(* Logix 5000 project; controller NWGG 1756-L72 rev 35.12; software revision 35.00; part 2 of 19 *)
(* tags used below, declared in another part *)
   T22 : TIMER[100];
   T4 : TIMER[100];

ADD_ON_INSTRUCTION Loadout_K_Valve_Control   (* revision 1.0 *)
VAR_IN_OUT
   K_Valve : udt_Loadout_K_Valve; {required}
   ALM_Clean_Pos_Failed : ALARM_DIGITAL; {required}
   ALM_Treat_Pos_Failed : ALARM_DIGITAL; {required}
   Treat_Position_Input : BOOL; {required}
   Clean_Position_Input : BOOL; {required}
   Clean_Gate_Relay : BOOL; {required}
   Treat_Gate_Relay : BOOL; {required}
END_VAR
VAR
   Clean_Pos_Failed_ACK : BOOL; {access None}
   Treat_Pos_Failedt_ACK : BOOL; {access None}
END_VAR

ROUTINE Logic   (* ladder *)
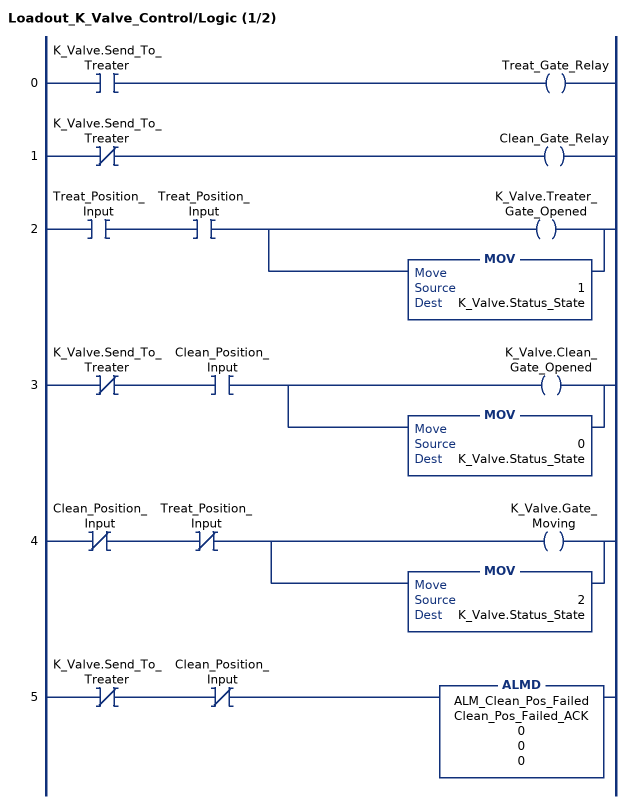
   0: XIC(K_Valve.Send_To_Treater)OTE(Treat_Gate_Relay);
   1: XIO(K_Valve.Send_To_Treater)OTE(Clean_Gate_Relay);
   2: XIC(Treat_Position_Input)XIC(Treat_Position_Input)[OTE(K_Valve.Treater_Gate_Opened) ,MOV(1,K_Valve.Status_State) ];
   3: XIO(K_Valve.Send_To_Treater)XIC(Clean_Position_Input)[OTE(K_Valve.Clean_Gate_Opened) ,MOV(0,K_Valve.Status_State) ];
   4: XIO(Clean_Position_Input)XIO(Treat_Position_Input)[OTE(K_Valve.Gate_Moving) ,MOV(2,K_Valve.Status_State) ];
   5: XIO(K_Valve.Send_To_Treater)XIO(Clean_Position_Input)ALMD(ALM_Clean_Pos_Failed,Clean_Pos_Failed_ACK,0,0,0);
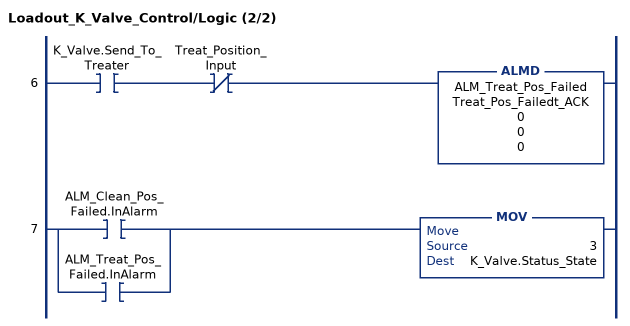
   6: XIC(K_Valve.Send_To_Treater)XIO(Treat_Position_Input)ALMD(ALM_Treat_Pos_Failed,Treat_Pos_Failedt_ACK,0,0,0);
   7: [XIC(ALM_Clean_Pos_Failed.InAlarm) ,XIC(ALM_Treat_Pos_Failed.InAlarm) ]MOV(3,K_Valve.Status_State);
END_ROUTINE
END_ADD_ON_INSTRUCTION

ADD_ON_INSTRUCTION Motor_Control   (* revision 1.0 *)
VAR_IN_OUT
   Motor_Contact : BOOL; {required}
END_VAR
VAR_INPUT
   Spd_20_Pct : BOOL; {required}
   Spd_10_Pct : BOOL; {required}
END_VAR
VAR_OUTPUT
   Running : BOOL; {access Read Only, required}
END_VAR
VAR_IN_OUT
   Motor_Alarm_SPD20 : ALARM_DIGITAL; {required}
   Motor_Alarm_SPD10 : ALARM_DIGITAL; {required}
   Motor_Alarm_Stopped_Over_Amps : ALARM_DIGITAL; {required}
   Motor_Start : udt_Motor_Start; {required}
END_VAR
VAR_INPUT
   Plugged_Sensor : BOOL; {required}
END_VAR
VAR_IN_OUT
   Motor_Alarm_Plugged : ALARM_DIGITAL; {required}
END_VAR
VAR_INPUT
   Motor_Amps : REAL; {required}
END_VAR
VAR_IN_OUT
   Motor_Config : udt_Motor_Config; {required}
   Motor_Starting : BOOL; {required}
   Motor_Alarm_Wont_Start : ALARM_DIGITAL; {required}
END_VAR
VAR_OUTPUT
   In_Alarm : BOOL; {access Read Only}
END_VAR
VAR_IN_OUT
   Treat_Batch_Status : DINT; {required}
   Clean_Batch_Status : DINT; {required}
   Transfer_Batch_Status : DINT; {required}
END_VAR
VAR_OUTPUT
   Motor_Batch_Ready : BOOL; {access Read Only}
END_VAR
VAR_IN_OUT
   Manual_Mode : BOOL; {required}
   InterLocked_Belt : BOOL; {required}
END_VAR
VAR_OUTPUT
   Motor_Batch_Ready_Clean : BOOL; {access Read Only}
   Motor_Batch_Ready_Treat : BOOL; {access Read Only}
   Motor_Batch_Ready_Transfer : BOOL; {access Read Only}
END_VAR
VAR
   TMR_BELT_SPD20 : TIMER := (PRE := 2000); {access None}
   TMR_AMP_INRUSH : TIMER := (PRE := 2000); {access None}
   Alm_Spd20_AK : BOOL; {access None}
   Alm_Spd10_AK : BOOL; {access None}
   Alm_Plugged_AK : BOOL; {access None}
   Alm_OVR_AMP_AK : BOOL; {access None}
   Stop_Motor_Plugged : BOOL; {access None}
   Stop_Motor_SLP20 : BOOL; {access None}
   Stop_Motor : BOOL; {access None}
   Stop_Motor_Ovr_Amp : BOOL; {access None}
   TMR_BELT_SPD10 : TIMER := (PRE := 2000); {access None}
   Alm_Wont_Start_AK : BOOL; {access None}
   Req_Motor_Start : BOOL; {access None}
   tmr_Auto_Stop_Delay : TIMER; {access None}
END_VAR

ROUTINE Logic   (* ladder *)
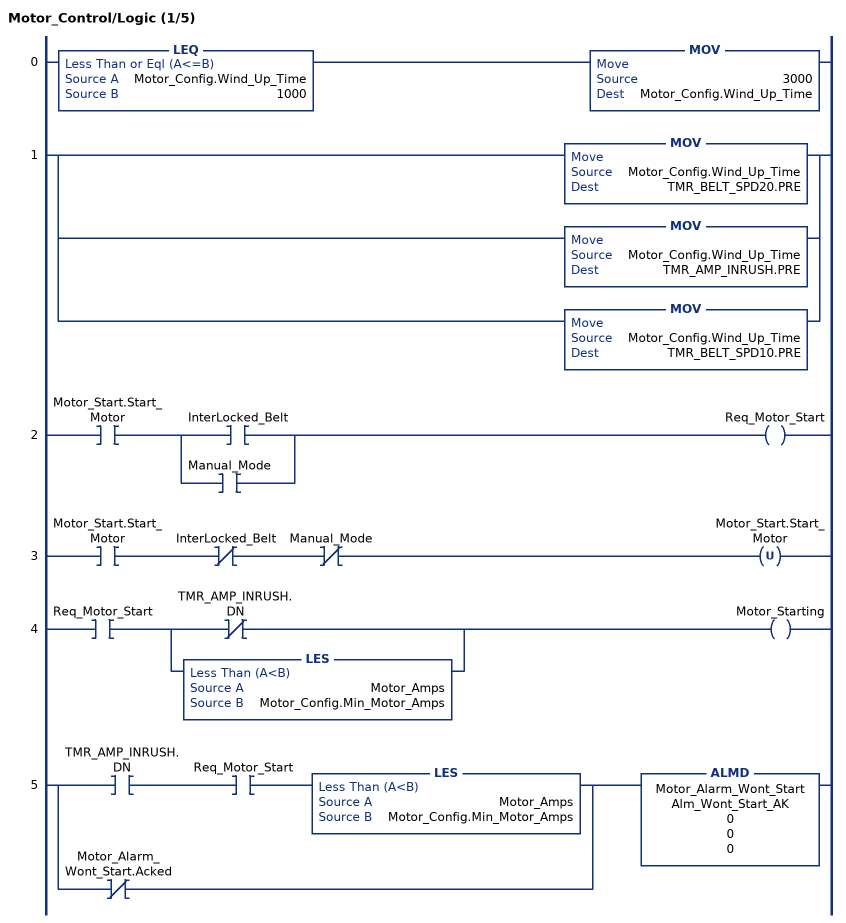
   0: LEQ(Motor_Config.Wind_Up_Time,1000)MOV(3000,Motor_Config.Wind_Up_Time);
   1: [MOV(Motor_Config.Wind_Up_Time,TMR_BELT_SPD20.PRE) ,MOV(Motor_Config.Wind_Up_Time,TMR_AMP_INRUSH.PRE) ,MOV(Motor_Config.Wind_Up_Time,TMR_BELT_SPD10.PRE) ];
   2: XIC(Motor_Start.Start_Motor)[XIC(InterLocked_Belt) ,XIC(Manual_Mode) ]OTE(Req_Motor_Start);
   3: XIC(Motor_Start.Start_Motor)XIO(InterLocked_Belt)XIO(Manual_Mode)OTU(Motor_Start.Start_Motor);
   4: XIC(Req_Motor_Start)[XIO(TMR_AMP_INRUSH.DN) ,LES(Motor_Amps,Motor_Config.Min_Motor_Amps) ]OTE(Motor_Starting);
   5: [XIC(TMR_AMP_INRUSH.DN) XIC(Req_Motor_Start) LES(Motor_Amps,Motor_Config.Min_Motor_Amps) ,XIO(Motor_Alarm_Wont_Start.Acked) ]ALMD(Motor_Alarm_Wont_Start,Alm_Wont_Start_AK,0,0,0);
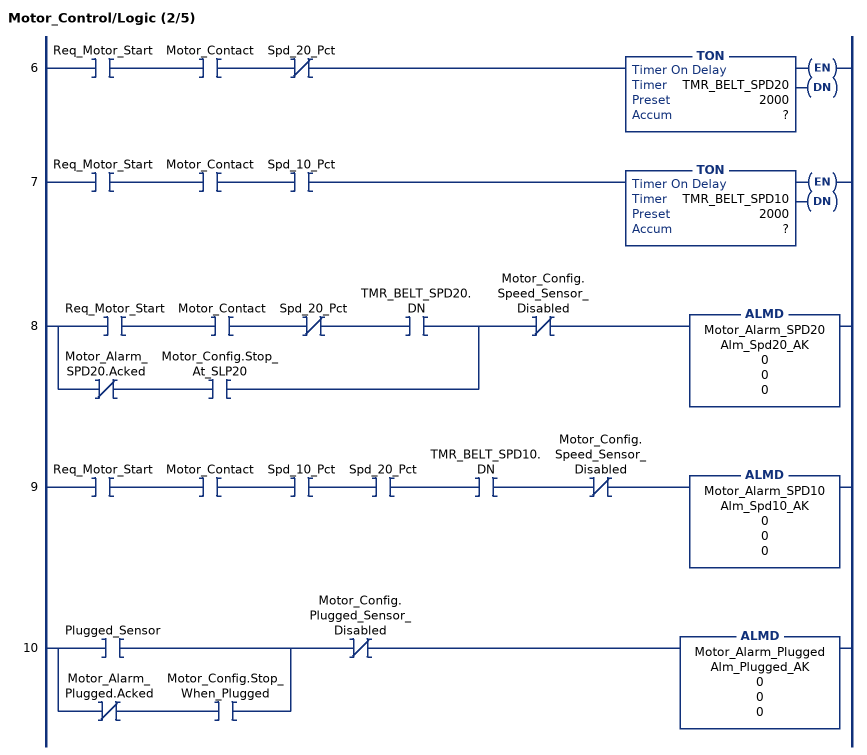
   6: XIC(Req_Motor_Start)XIC(Motor_Contact)XIO(Spd_20_Pct)TON(TMR_BELT_SPD20,?,?);
   7: XIC(Req_Motor_Start)XIC(Motor_Contact)XIC(Spd_10_Pct)TON(TMR_BELT_SPD10,?,?);
   8: [XIC(Req_Motor_Start) XIC(Motor_Contact) XIO(Spd_20_Pct) XIC(TMR_BELT_SPD20.DN) ,XIO(Motor_Alarm_SPD20.Acked) XIC(Motor_Config.Stop_At_SLP20) ]XIO(Motor_Config.Speed_Sensor_Disabled)ALMD(Motor_Alarm_SPD20,Alm_Spd20_AK,0,0,0);
   9: XIC(Req_Motor_Start)XIC(Motor_Contact)XIC(Spd_10_Pct)XIC(Spd_20_Pct)XIC(TMR_BELT_SPD10.DN)XIO(Motor_Config.Speed_Sensor_Disabled)ALMD(Motor_Alarm_SPD10,Alm_Spd10_AK,0,0,0);
   10: [XIC(Plugged_Sensor) ,XIO(Motor_Alarm_Plugged.Acked) XIC(Motor_Config.Stop_When_Plugged) ]XIO(Motor_Config.Plugged_Sensor_Disabled)ALMD(Motor_Alarm_Plugged,Alm_Plugged_AK,0,0,0);
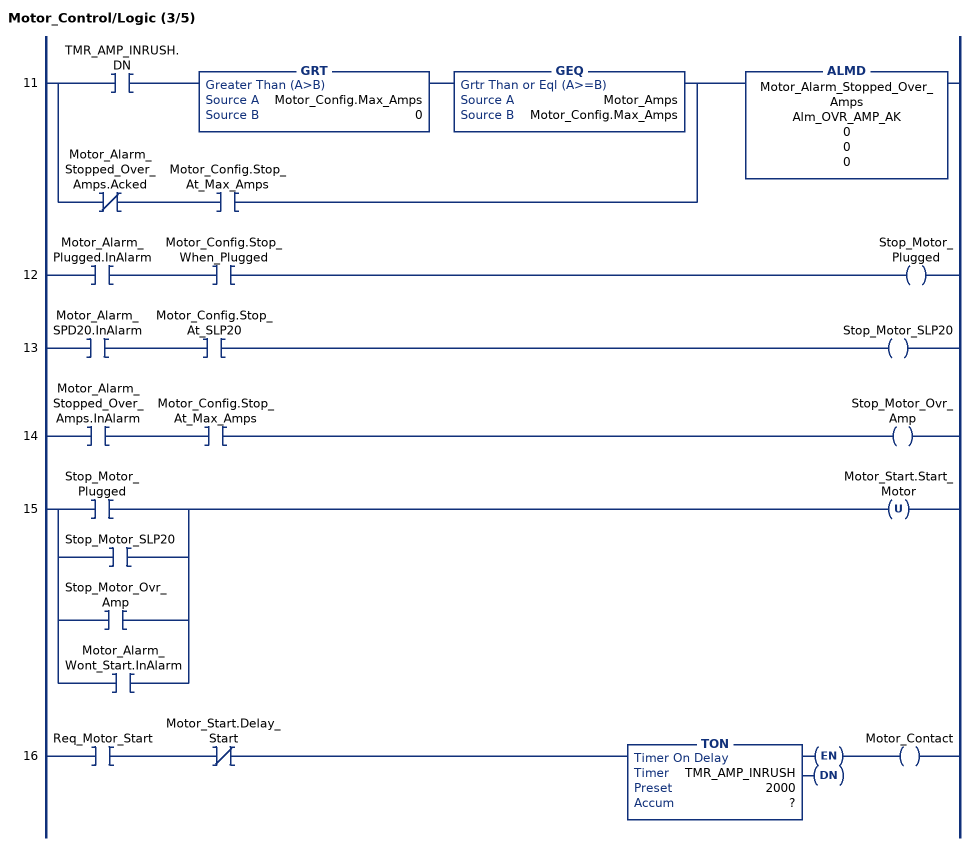
   11: [XIC(TMR_AMP_INRUSH.DN) GRT(Motor_Config.Max_Amps,0) GEQ(Motor_Amps,Motor_Config.Max_Amps) ,XIO(Motor_Alarm_Stopped_Over_Amps.Acked) XIC(Motor_Config.Stop_At_Max_Amps) ]ALMD(Motor_Alarm_Stopped_Over_Amps,Alm_OVR_AMP_AK,0,0,0);
   12: XIC(Motor_Alarm_Plugged.InAlarm)XIC(Motor_Config.Stop_When_Plugged)OTE(Stop_Motor_Plugged);
   13: XIC(Motor_Alarm_SPD20.InAlarm)XIC(Motor_Config.Stop_At_SLP20)OTE(Stop_Motor_SLP20);
   14: XIC(Motor_Alarm_Stopped_Over_Amps.InAlarm)XIC(Motor_Config.Stop_At_Max_Amps)OTE(Stop_Motor_Ovr_Amp);
   15: [XIC(Stop_Motor_Plugged) ,XIC(Stop_Motor_SLP20) ,XIC(Stop_Motor_Ovr_Amp) ,XIC(Motor_Alarm_Wont_Start.InAlarm) ]OTU(Motor_Start.Start_Motor);
   16: XIC(Req_Motor_Start)XIO(Motor_Start.Delay_Start)TON(TMR_AMP_INRUSH,?,?)OTE(Motor_Contact);
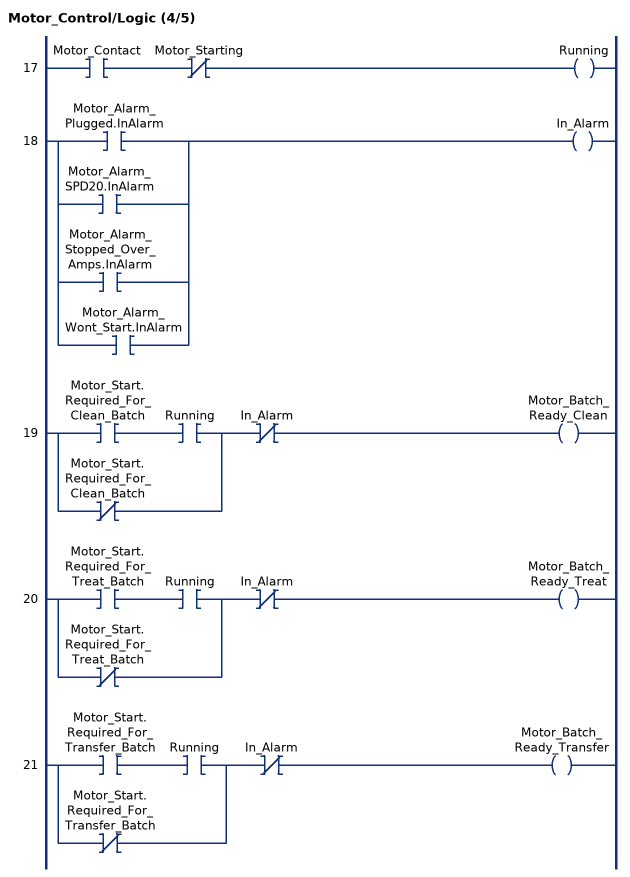
   17: XIC(Motor_Contact)XIO(Motor_Starting)OTE(Running);
   18: [XIC(Motor_Alarm_Plugged.InAlarm) ,XIC(Motor_Alarm_SPD20.InAlarm) ,XIC(Motor_Alarm_Stopped_Over_Amps.InAlarm) ,XIC(Motor_Alarm_Wont_Start.InAlarm) ]OTE(In_Alarm);
   19: [XIC(Motor_Start.Required_For_Clean_Batch) XIC(Running) ,XIO(Motor_Start.Required_For_Clean_Batch) ]XIO(In_Alarm)OTE(Motor_Batch_Ready_Clean);
   20: [XIC(Motor_Start.Required_For_Treat_Batch) XIC(Running) ,XIO(Motor_Start.Required_For_Treat_Batch) ]XIO(In_Alarm)OTE(Motor_Batch_Ready_Treat);
   21: [XIC(Motor_Start.Required_For_Transfer_Batch) XIC(Running) ,XIO(Motor_Start.Required_For_Transfer_Batch) ]XIO(In_Alarm)OTE(Motor_Batch_Ready_Transfer);
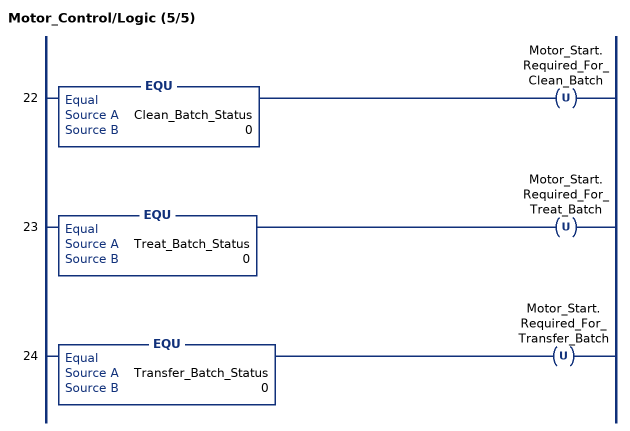
   22: EQU(Clean_Batch_Status,0)OTU(Motor_Start.Required_For_Clean_Batch);
   23: EQU(Treat_Batch_Status,0)OTU(Motor_Start.Required_For_Treat_Batch);
   24: EQU(Transfer_Batch_Status,0)OTU(Motor_Start.Required_For_Transfer_Batch);
END_ROUTINE
END_ADD_ON_INSTRUCTION

ADD_ON_INSTRUCTION SCP   (* revision 1.0, vendor Rockwell Automation *)
VAR_INPUT
   In : ALIAS FOR SCL_01.In; {access None, required}
   InRawMin : REAL; {access None, required}
   InRawMax : REAL; {required}
   InEUMin : REAL; {required}
   InEUMax : REAL; {required}
   Out : DINT; {required}
END_VAR
VAR
   SCL_01 : SCALE; {access None}
   SUB_01 : FBD_MATH; {access None}
   SEL_01 : SELECT; {access None}
   SCL_02 : SCALE; {access None}
   LES_02 : FBD_COMPARE; {access None}
   __l56AFB0E5191E6558 : REAL; {access None}
   __l0BF49CB3D0F7F241 : REAL; {access None}
   __l7339031870541241 : REAL; {access None}
   __l88E0968931849F84 : REAL; {access None}
END_VAR

ROUTINE Logic   (* function block diagram *)
   SHEET 1
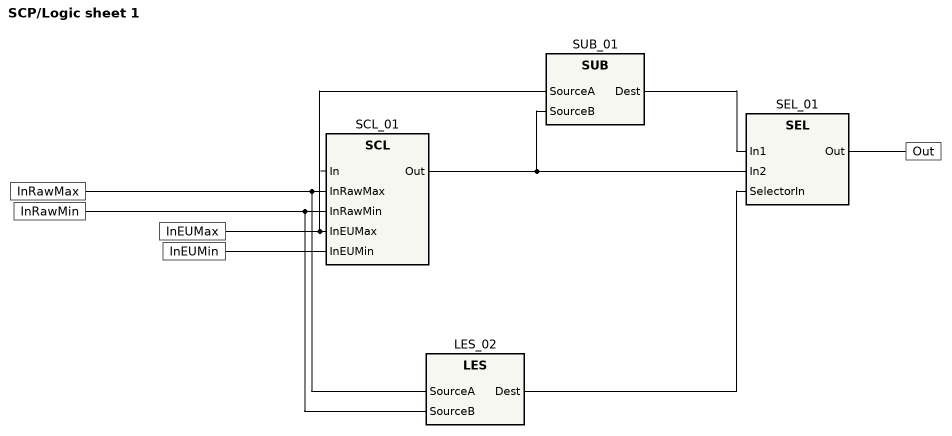
   SCL_01 : SCL(InRawMax := InRawMax, InRawMin := InRawMin, InEUMax := InEUMax, InEUMin := InEUMin);   // unwired pins: In
   LES_02 : LES(SourceA := InRawMax, SourceB := InRawMin);
   SUB_01 : SUB(SourceA := InEUMax, SourceB := SCL_01.Out);
   SEL_01 : SEL(In1 := SUB_01.Dest, In2 := SCL_01.Out, SelectorIn := LES_02.Dest);
   Out := SEL_01.Out;
END_ROUTINE
END_ADD_ON_INSTRUCTION

ADD_ON_INSTRUCTION SCP_Inv   (* revision 1.0, vendor Rockwell Automation *)
VAR_INPUT
   In : ALIAS FOR SCL_01.In; {access None, required}
   InRawMin : REAL; {access None, required}
   InRawMax : REAL; {required}
   InEUMin : REAL; {required}
   InEUMax : REAL; {required}
END_VAR
VAR_OUTPUT
   Out : REAL; {required}
END_VAR
VAR
   SCL_01 : SCALE; {access None}
   SUB_01 : FBD_MATH; {access None}
   SEL_01 : SELECT; {access None}
   SCL_02 : SCALE; {access None}
   LES_02 : FBD_COMPARE; {access None}
   __lC7D96F2B3EA1267C : REAL; {access None}
   __lD4FD1BAAF7FBA06E : REAL; {access None}
   __lFFF49F1C0E6A2B2A : REAL; {access None}
   __lEB05C44F0520614F : REAL; {access None}
END_VAR

ROUTINE Logic   (* function block diagram *)
   SHEET 1
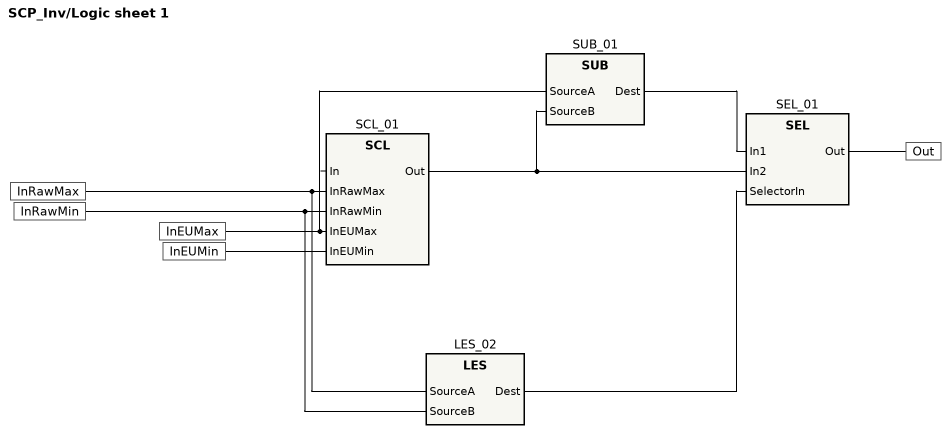
   SCL_01 : SCL(InRawMax := InRawMax, InRawMin := InRawMin, InEUMax := InEUMax, InEUMin := InEUMin);   // unwired pins: In
   LES_02 : LES(SourceA := InRawMax, SourceB := InRawMin);
   SUB_01 : SUB(SourceA := InEUMax, SourceB := SCL_01.Out);
   SEL_01 : SEL(In1 := SUB_01.Dest, In2 := SCL_01.Out, SelectorIn := LES_02.Dest);
   Out := SEL_01.Out;
END_ROUTINE
END_ADD_ON_INSTRUCTION

ADD_ON_INSTRUCTION Truck_Scale_Control   (* revision 1.0 *)
VAR_IN_OUT
   Scale : udt_Truck_Scale; {required}
   Scale_Output : AB:ETHERNET_MODULE_DINT_4Bytes:O:0; {required}
   Scale_Input : AB:ETHERNET_MODULE_DINT_4Bytes:I:0; {required}
END_VAR
VAR
   Rate_Tmr : TIMER := (PRE := 1000, ACC := 713); {access None}
   Accum_Rate_Index1 : COUNTER := (PRE := 11); {access None}
   Old_Accum_Rate : REAL; {access None}
   Rate_Tare : REAL; {access None}
   Lock_Stable_Rate : DINT; {access None}
   Scale_Avg1 : REAL[15]; {access None}
   tmr_Stable : TIMER := (PRE := 2000); {access None}
   tmr_Old_Rate : TIMER := (PRE := 1000); {access None}
   Scale_Avg2 : REAL[15]; {access None}
   Scale_Avg3 : REAL[15]; {access None}
   Avg_Rate1 : REAL; {access None}
   Avg_Rate2 : REAL; {access None}
   Accum_Rate_Index2 : COUNTER := (PRE := 5); {access None}
   Accum_Rate_Index3 : COUNTER := (PRE := 5); {access None}
   Avg_Rate3 : DINT; {access None}
   tmrWeightTest : TIMER; {access None}
END_VAR

ROUTINE Logic   (* ladder *)
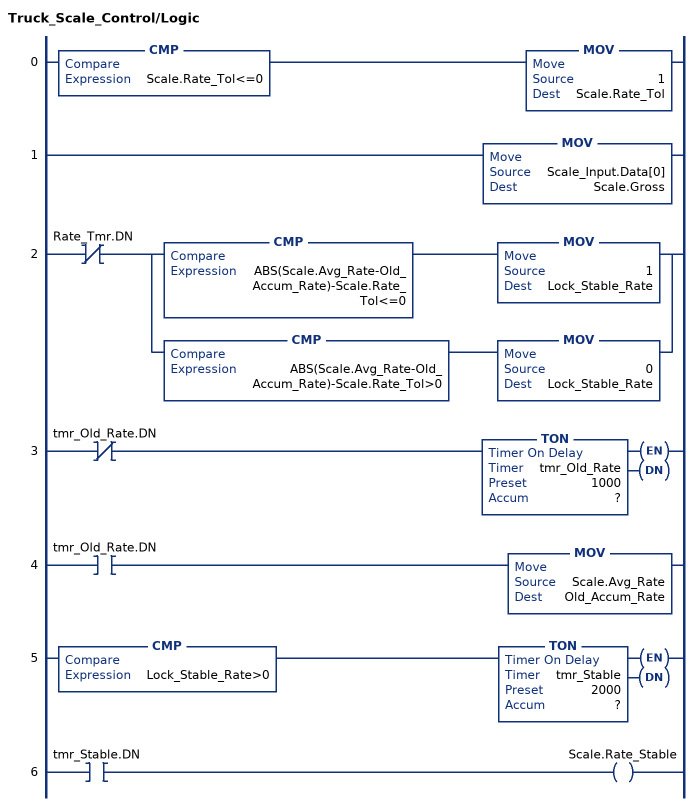
   0: CMP(Scale.Rate_Tol<=0)MOV(1,Scale.Rate_Tol);
   1: MOV(Scale_Input.Data[0],Scale.Gross);
   2: XIO(Rate_Tmr.DN)[CMP(ABS(Scale.Avg_Rate-Old_Accum_Rate)-Scale.Rate_Tol<=0) MOV(1,Lock_Stable_Rate) ,CMP(ABS(Scale.Avg_Rate-Old_Accum_Rate)-Scale.Rate_Tol>0) MOV(0,Lock_Stable_Rate) ];
   3: XIO(tmr_Old_Rate.DN)TON(tmr_Old_Rate,?,?);
   4: XIC(tmr_Old_Rate.DN)MOV(Scale.Avg_Rate,Old_Accum_Rate);
   5: CMP(Lock_Stable_Rate>0)TON(tmr_Stable,?,?);
   6: XIC(tmr_Stable.DN)OTE(Scale.Rate_Stable);
END_ROUTINE
END_ADD_ON_INSTRUCTION

VAR_GLOBAL   (* controller tags *)
   _100AUTO : ALIAS FOR B9[100].4;
   _100HAND : ALIAS FOR B9[100].3;
   _100MB : ALIAS FOR B9[100].2;
   _100STB : ALIAS FOR B9[100].0;
   _100STPB : ALIAS FOR B9[100].1;
   _101_FEED_AUGER_PIT_101_HM : HOUR_METER := (HR_METER_DISPLAY := 21700, MAINTENANCE_ALARM := 1);
   _101AUTO : ALIAS FOR B9[101].4;
   _101HAND : ALIAS FOR B9[101].3;
   _101M : ALIAS FOR O25[9].3;
   _101MB : ALIAS FOR B9[101].2;
   _101STB : ALIAS FOR B9[101].0;
   _101STPB : ALIAS FOR B9[101].1;
   _101Y : ALIAS FOR I25[1].3;
   _102_EXPLORE_TANK_41_RECEIVING_LEG_HM : HOUR_METER := (MOTOR_RUNNING_INPUT_1 := 1, HR_METER_DISPLAY := 13009, MAINTENANCE_ALARM := 1);
   _102AUTO : ALIAS FOR B9[102].4;
   _102HAND : ALIAS FOR B9[102].3;
   _102M : ALIAS FOR O25[8].9;
   _102MB : ALIAS FOR B9[102].2;
   _102STB : ALIAS FOR B9[102].0;
   _102STPB : ALIAS FOR B9[102].1;
   _102Y : ALIAS FOR I25[0].9;
   _103_TANK_42_RECEIVING_LEG_HM : HOUR_METER := (HR_METER_DISPLAY := 4431, NEXT_SCHDL_MAINTENANCE := 2, MAINTENANCE_ALARM := 1);
   _103_TANK_42_RECEIVING_LEG_RUNNING : BOOL;
   _103AUTO : ALIAS FOR B9[103].4;
   _103HAND : ALIAS FOR B9[103].3;
   _103M : ALIAS FOR O25[8].12;
   _103MB : ALIAS FOR B9[103].2;
   _103STB : ALIAS FOR B9[103].0;
   _103STPB : ALIAS FOR B9[103].1;
   _103Y : ALIAS FOR I25[0].12;
   _106_TANK_17_AUGER_HM : HOUR_METER := (HR_METER_DISPLAY := 5679, NEXT_SCHDL_MAINTENANCE := 2, MAINTENANCE_ALARM := 1);
   _106_TANK_17_AUGER_RUNNING : BOOL;
   _106AUTO : ALIAS FOR B9[106].4;
   _106HAND : ALIAS FOR B9[106].3;
   _106M : ALIAS FOR O25[9].5;
   _106MB : ALIAS FOR B9[106].2;
   _106STB : ALIAS FOR B9[106].0;
   _106STPB : ALIAS FOR B9[106].1;
   _106Y : ALIAS FOR I25[1].5;
   _107_SOUTH_BELT_HM : HOUR_METER := (MOTOR_RUNNING_INPUT_1 := 1, HR_METER_DISPLAY := 11100, NEXT_SCHDL_MAINTENANCE := 2, MAINTENANCE_ALARM := 1);
   _107_TANKS_1THRU7_SOUTH_RUNNING : BOOL := 1;
   _107AUTO : ALIAS FOR B9[107].4;
   _107HAND : ALIAS FOR B9[107].3;
   _107M : ALIAS FOR O25[9].12;
   _107MB : ALIAS FOR B9[107].2;
   _107PS : ALIAS FOR I25[4].2;
   _107PSB : ALIAS FOR B9[107].5;
   _107STB : ALIAS FOR B9[107].0;
   _107STPB : ALIAS FOR B9[107].1;
   _107Y : ALIAS FOR I25[1].12;
   _108_CENTER_BELT_HM : HOUR_METER := (MOTOR_RUNNING_INPUT_1 := 1, HR_METER_DISPLAY := 19687, NEXT_SCHDL_MAINTENANCE := 2, MAINTENANCE_ALARM := 1);
   _108_CENTER_BELT_RUNNING : BOOL := 1;
   _108AUTO : ALIAS FOR B9[108].4;
   _108HAND : ALIAS FOR B9[108].3;
   _108M : ALIAS FOR O25[10].15;
   _108MB : ALIAS FOR B9[108].2;
   _108PS : ALIAS FOR I25[4].1;
   _108STB : ALIAS FOR B9[108].0;
   _108STPB : ALIAS FOR B9[108].1;
   _108Y : ALIAS FOR I25[2].15;
   _109_NORTH_BELT_HM : HOUR_METER := (HR_METER_DISPLAY := 77, NEXT_SCHDL_MAINTENANCE := 2, MAINTENANCE_ALARM := 1);
   _109_PS_DLY : ALIAS FOR T11[4];
   _109_RAW_RECEIVING_NORTH_BELT_RUNNING : BOOL;
   _109_SLOW_D : ALIAS FOR T11[5];
   _109_SLW_SP : ALIAS FOR I25[3].14;
   _109_STOP_D : ALIAS FOR T11[6];
   _109_STP_SP : ALIAS FOR I25[3].15;
   _109AUTO : ALIAS FOR B9[109].4;
   _109HAND : ALIAS FOR B9[109].3;
   _109M : ALIAS FOR O25[10].9;
   _109MB : ALIAS FOR B9[109].2;
   _109PS : ALIAS FOR I25[4].0;
   _109STB : ALIAS FOR B9[109].0;
   _109STPB : ALIAS FOR B9[109].1;
   _109Y : ALIAS FOR I25[2].9;
   _10AUTO : ALIAS FOR B9[10].4;
   _10HAND : ALIAS FOR B9[10].3;
   _10MB : ALIAS FOR B9[10].2;
   _10STB : ALIAS FOR B9[10].0;
   _10STPB : ALIAS FOR B9[10].1;
   _10Y : ALIAS FOR I25[0].11;
   _110_TANK_16_AUGER_HM : HOUR_METER := (HR_METER_DISPLAY := 3779, NEXT_SCHDL_MAINTENANCE := 2, MAINTENANCE_ALARM := 1);
   _110_TANK_16_AUGER_RUNNING : BOOL;
   _110AUTO : ALIAS FOR B9[110].4;
   _110HAND : ALIAS FOR B9[110].3;
   _110M : ALIAS FOR O25[8].15;
   _110MB : ALIAS FOR B9[110].2;
   _110STB : ALIAS FOR B9[110].0;
   _110STPB : ALIAS FOR B9[110].1;
   _110Y : ALIAS FOR I25[0].15;
   _111_TANK_17_AUGER_HM : HOUR_METER := (HR_METER_DISPLAY := 1055, MAINTENANCE_ALARM := 1);
   _111AUTO : ALIAS FOR B9[111].4;
   _111HAND : ALIAS FOR B9[111].3;
   _111M : ALIAS FOR O25[9].0;
   _111MB : ALIAS FOR B9[111].2;
   _111STB : ALIAS FOR B9[111].0;
   _111STPB : ALIAS FOR B9[111].1;
   _111Y : ALIAS FOR I25[1].0;
   _113_GATE_B : ALIAS FOR I25[4].12;
   _113_GATE_B1 : ALIAS FOR I25[4].13;
   _113_HIGHROLLER_TANKS_11TO15_HM : HOUR_METER := (HR_METER_DISPLAY := 1063, NEXT_SCHDL_MAINTENANCE := 2, MAINTENANCE_ALARM := 1);
   _113_HIGHROLLER_TANKS_11TO15_RUNNING : BOOL;
   _113_TO_BC1 : ALIAS FOR O25[11].9;
   _113_TO_BC9 : ALIAS FOR O25[11].8;
   _113AUTO : ALIAS FOR B9[113].4;
   _113HAND : ALIAS FOR B9[113].3;
   _113M : ALIAS FOR O25[10].5;
   _113MB : ALIAS FOR B9[113].2;
   _113STB : ALIAS FOR B9[113].0;
   _113STPB : ALIAS FOR B9[113].1;
   _113Y : ALIAS FOR I25[2].5;
   _114_TANKS_1THRU7_NORTH_HM : HOUR_METER := (HR_METER_DISPLAY := 9528, MAINTENANCE_ALARM := 1);
   _114_TANKS_1THRU7_NORTH_RUNNING : BOOL;
   _115_M : ALIAS FOR O25[22].0;
   _115AUTO : ALIAS FOR B9[115].4;
   _115HAND : ALIAS FOR B9[115].3;
   _115MB : ALIAS FOR B9[115].2;
   _115STB : ALIAS FOR B9[115].0;
   _115STPB : ALIAS FOR B9[115].1;
   _116_DRAG_16_HM : HOUR_METER := (HR_METER_DISPLAY := 3781, MAINTENANCE_ALARM := 1);
   _116AUTO : ALIAS FOR B9[116].4;
   _116HAND : ALIAS FOR B9[116].3;
   _116M : ALIAS FOR O25[10].10;
   _116MB : ALIAS FOR B9[116].2;
   _116STB : ALIAS FOR B9[116].0;
   _116STPB : ALIAS FOR B9[116].1;
   _116Y : ALIAS FOR I25[2].10;
   _117_DRAG_17_HM : HOUR_METER := (HR_METER_DISPLAY := 5681, MAINTENANCE_ALARM := 1);
   _117AUTO : ALIAS FOR B9[117].4;
   _117HAND : ALIAS FOR B9[117].3;
   _117M : ALIAS FOR O25[10].8;
   _117MB : ALIAS FOR B9[117].2;
   _117STB : ALIAS FOR B9[117].0;
   _117STPB : ALIAS FOR B9[117].1;
   _117Y : ALIAS FOR I25[2].8;
   _11_BINDICA : ALIAS FOR B15[11].0;
   _11_BINDICA1 : ALIAS FOR B15[11].1;
   _11_GATE_PO : ALIAS FOR I16[0];
   _11_GATE_PO1 : ALIAS FOR N14[11];
   _11_GATE_PO_STOR : REAL := 86.33458;
   _11_PS : ALIAS FOR I25[4].14;
   _11_PS_DLY : ALIAS FOR T11[2];
   _11_SLOW_SP : ALIAS FOR I25[4].3;
   _11_STOP_SP : ALIAS FOR I25[4].6;
   _11_TANK_41_42_HIGHROLLER_HM : HOUR_METER := (HR_METER_DISPLAY := 6844, NEXT_SCHDL_MAINTENANCE := 2, MAINTENANCE_ALARM := 1);
   _11_TANK_41_42_HIGHROLLER_RUNNING : BOOL;
   _11_VALVE_R : ALIAS FOR I25[4].4;
   _11_VALVE_S : ALIAS FOR I25[4].5;
   _11AUTO : ALIAS FOR B9[11].4;
   _11HAND : ALIAS FOR B9[11].3;
   _11M : ALIAS FOR O25[9].2;
   _11MB : ALIAS FOR B9[11].2;
   _11STB : ALIAS FOR B9[11].0;
   _11STPB : ALIAS FOR B9[11].1;
   _11Y : ALIAS FOR I25[1].2;
   _122_RECIEVING_LEG_HM : HOUR_METER := (MOTOR_RUNNING_INPUT_1 := 1, HR_METER_DISPLAY := 24537, MAINTENANCE_ALARM := 1);
   _122AUTO : ALIAS FOR B9[122].4;
   _122HAND : ALIAS FOR B9[122].3;
   _122M : ALIAS FOR O25[9].1;
   _122MB : ALIAS FOR B9[122].2;
   _122STB : ALIAS FOR B9[122].0;
   _122STPB : ALIAS FOR B9[122].1;
   _122Y : ALIAS FOR I25[1].1;
   _123_CLEAN_LEG_HM : HOUR_METER := (MOTOR_RUNNING_INPUT_1 := 1, HR_METER_DISPLAY := 26622, NEXT_SCHDL_MAINTENANCE := 2, MAINTENANCE_ALARM := 1);
   _123_CLEAN_LEG_RUNNING : BOOL := 1;
   _123_COMPUW : ALIAS FOR I18[7];
   _123_COMPUW1 : ALIAS FOR N7[20];
   _123AUTO : ALIAS FOR B9[123].4;
   _123HAND : ALIAS FOR B9[123].3;
   _123M : ALIAS FOR O25[10].6;
   _123MB : ALIAS FOR B9[123].2;
   _123STB : ALIAS FOR B9[123].0;
   _123STPB : ALIAS FOR B9[123].1;
   _123Y : ALIAS FOR I25[2].6;
   _124AUTO : ALIAS FOR B9[124].4;
   _124HAND : ALIAS FOR B9[124].3;
   _124M : ALIAS FOR O25[9].13;
   _124MB : ALIAS FOR B9[124].2;
   _124STB : ALIAS FOR B9[124].0;
   _124STPB : ALIAS FOR B9[124].1;
   _125_COLOR_SORTER_LEG_HM : HOUR_METER := (MOTOR_RUNNING_INPUT_1 := 1, HR_METER_DISPLAY := 26513, NEXT_SCHDL_MAINTENANCE := 2, MAINTENANCE_ALARM := 1);
   _126_ASPERATOR : HOUR_METER := (MOTOR_RUNNING_INPUT_1 := 1, HR_METER_DISPLAY := 25758, NEXT_SCHDL_MAINTENANCE := 2, MAINTENANCE_ALARM := 1);
   _128_SCREENINGS_DRAG_HM : HOUR_METER := (MOTOR_RUNNING_INPUT_1 := 1, HR_METER_DISPLAY := 26532, NEXT_SCHDL_MAINTENANCE := 2, MAINTENANCE_ALARM := 1);
   _12_BINDICA : ALIAS FOR B15[12].0;
   _12_BINDICA1 : ALIAS FOR B15[12].1;
   _12_GATE_PO : ALIAS FOR I16[1];
   _12_GATE_PO1 : ALIAS FOR N14[12];
   _12_GATE_PO_STOR : REAL := 94.72872;
   _13_BINDICA : ALIAS FOR B15[13].0;
   _13_BINDICA1 : ALIAS FOR B15[13].1;
   _13_GATE_PO : ALIAS FOR I16[2];
   _13_GATE_PO1 : ALIAS FOR N14[13];
   _13_GATE_PO_STOR : REAL := 79.42468;
   _14_BINDICA : ALIAS FOR B15[14].0;
   _14_BINDICA1 : ALIAS FOR B15[14].1;
   _14_GATE_PO : ALIAS FOR I16[3];
   _14_GATE_PO1 : ALIAS FOR N14[14];
   _14_GATE_PO_STOR : REAL := 93.90426;
   _15_BINDICA : ALIAS FOR B15[15].0;
   _15_BINDICA1 : ALIAS FOR B15[15].1;
   _15_GATE_PO : ALIAS FOR I16[4];
   _15_GATE_PO1 : ALIAS FOR N14[15];
   _15_GATE_PO_STOR : REAL := 92.96653;
   _16_BINDICA : ALIAS FOR B15[16].0;
   _16_BINDICA1 : ALIAS FOR B15[16].1;
   _16_GATE_PO : ALIAS FOR I16[5];
   _16_GATE_PO1 : ALIAS FOR N14[16];
   _16_GATE_PO_STOR : REAL := 30.742159;
   _17_BINDICA : ALIAS FOR B15[17].0;
   _17_BINDICA1 : ALIAS FOR B15[17].1;
   _17_GATE_PO : ALIAS FOR I16[6];
   _17_GATE_PO1 : ALIAS FOR N14[17];
   _17_GATE_PO_STOR : REAL := 78.57861;
   _1_CLEAN_SEED_UPPER_BELT_HM : HOUR_METER := (MOTOR_RUNNING_INPUT_1 := 1, HR_METER_DISPLAY := 13589, NEXT_SCHDL_MAINTENANCE := 2, MAINTENANCE_ALARM := 1);
   _1_CLEAN_SEED_UPPER_BELT_RUNNING : BOOL := 1;
   _1AUTO : ALIAS FOR B9[1].4;
   _1HAND : ALIAS FOR B9[1].3;
   _1M : ALIAS FOR O25[9].8;
   _1MB : ALIAS FOR B9[1].2;
   _1STB : ALIAS FOR B9[1].0;
   _1STPB : ALIAS FOR B9[1].1;
   _1Y : ALIAS FOR I25[1].8;
   _21_BINDICA : ALIAS FOR B15[21].0;
   _21_BINDICA1 : ALIAS FOR B15[21].1;
   _21_GATE_PO : ALIAS FOR I16[7];
   _21_GATE_PO1 : ALIAS FOR N14[21];
   _21_GATE_PO_STOR : REAL := 87.275024;
   _22_BINDICA : ALIAS FOR B15[22].0;
   _22_BINDICA1 : ALIAS FOR B15[22].1;
   _22_GATE_PO : ALIAS FOR I17[0];
   _22_GATE_PO1 : ALIAS FOR N14[22];
   _22_GATE_PO_STOR : REAL := 83.08857;
   _22AUTO : ALIAS FOR B9[22].4;
   _22HAND : ALIAS FOR B9[22].3;
   _22MB : ALIAS FOR B9[22].2;
   _22STB : ALIAS FOR B9[22].0;
   _22STPB : ALIAS FOR B9[22].1;
   _23_BINDICA : ALIAS FOR B15[23].0;
   _23_BINDICA1 : ALIAS FOR B15[23].1;
   _23_GATE_PO : ALIAS FOR I17[1];
   _23_GATE_PO1 : ALIAS FOR N14[23];
   _23_GATE_PO_STOR : REAL := 96.74677;
   _24_16_0 : ALIAS FOR N250[0];
   _24_16_1 : ALIAS FOR N250[1];
   _24_16_2 : ALIAS FOR N250[2];
   _24_16_3 : ALIAS FOR N250[3];
   _24_16_4 : ALIAS FOR N250[4];
   _24_16_5 : ALIAS FOR N250[5];
   _24_16_6 : ALIAS FOR N250[6];
   _24_16_7 : ALIAS FOR N250[7];
   _24_16_BLK : ALIAS FOR T4[58];
   _24_17_0 : ALIAS FOR N240[0];
   _24_17_1 : ALIAS FOR N240[1];
   _24_17_2 : ALIAS FOR N240[2];
   _24_17_3 : ALIAS FOR N240[3];
   _24_17_4 : ALIAS FOR N240[4];
   _24_17_5 : ALIAS FOR N240[5];
   _24_17_6 : ALIAS FOR N240[6];
   _24_17_7 : ALIAS FOR N240[7];
   _24_17_BLK : ALIAS FOR T4[57];
   _24_18_0_AN : ALIAS FOR N230[10];
   _24_18_1_AN : ALIAS FOR N230[11];
   _24_18_2_AN : ALIAS FOR N230[12];
   _24_18_3_AN : ALIAS FOR N230[13];
   _24_18_BLK : ALIAS FOR T4[40];
   _24_18_MULT : ALIAS FOR N230[14];
   _24_19_0 : ALIAS FOR N220[10];
   _24_19_1 : ALIAS FOR N220[11];
   _24_19_2 : ALIAS FOR N220[12];
   _24_19_3 : ALIAS FOR N220[13];
   _24_19_BLK : ALIAS FOR T4[39];
   _24_20_0 : ALIAS FOR N210[10];
   _24_20_1 : ALIAS FOR N210[11];
   _24_20_2 : ALIAS FOR N210[12];
   _24_20_3 : ALIAS FOR N210[13];
   _24_20_BLK : ALIAS FOR T4[38];
   _24_BINDICA : ALIAS FOR B15[24].0;
   _24_BINDICA1 : ALIAS FOR B15[24].1;
   _24_GATE_PO : ALIAS FOR I17[2];
   _24_GATE_PO1 : ALIAS FOR N14[24];
   _24_GATE_PO_STOR : REAL := 90.36168;
   _25_16_0 : ALIAS FOR N200[10];
   _25_16_1 : ALIAS FOR N200[11];
   _25_16_2 : ALIAS FOR N200[12];
   _25_16_3 : ALIAS FOR N200[13];
   _25_16_BLK : ALIAS FOR T4[37];
   _25_17_0 : ALIAS FOR N190[0];
   _25_17_1 : ALIAS FOR N190[1];
   _25_17_2 : ALIAS FOR N190[2];
   _25_17_3 : ALIAS FOR N190[3];
   _25_17_BLK : ALIAS FOR T4[36];
   _25_18_TMR : ALIAS FOR T4[35];
   _25_BINDICA : ALIAS FOR B15[25].0;
   _25_BINDICA1 : ALIAS FOR B15[25].1;
   _25_GATE_PO : ALIAS FOR I17[3];
   _25_GATE_PO1 : ALIAS FOR N14[25];
   _25_GATE_PO_STOR : REAL := 103.03115;
   _26_BINDICA : ALIAS FOR B15[26].0;
   _26_BINDICA1 : ALIAS FOR B15[26].1;
   _26_GATE_PO : ALIAS FOR I17[4];
   _26_GATE_PO1 : ALIAS FOR N14[26];
   _26_GATE_PO_STOR : REAL := 98.9571;
   _27_BINDICA : ALIAS FOR B15[27].0;
   _27_BINDICA1 : ALIAS FOR B15[27].1;
   _27_GATE_PO : ALIAS FOR I17[5];
   _27_GATE_PO1 : ALIAS FOR N14[27];
   _28_BINDICA : ALIAS FOR B15[28].0;
   _28_BINDICA1 : ALIAS FOR B15[28].1;
   _28_GATE_PO : ALIAS FOR I17[6];
   _28_GATE_PO1 : ALIAS FOR N14[28];
   _29_BINDICA : ALIAS FOR B15[29].0;
   _29_BINDICA1 : ALIAS FOR B15[29].1;
   _29_GATE_PO : ALIAS FOR I17[7];
   _29_GATE_PO1 : ALIAS FOR N14[29];
   _2AUTO : ALIAS FOR B9[2].4;
   _2HAND : ALIAS FOR B9[2].3;
   _2M : ALIAS FOR O25[9].15;
   _2MB : ALIAS FOR B9[2].2;
   _2STB : ALIAS FOR B9[2].0;
   _2STPB : ALIAS FOR B9[2].1;
   _2Y : ALIAS FOR I25[1].15;
   _35_JUMP_LEG_HM : HOUR_METER := (MOTOR_RUNNING_INPUT_1 := 1, HR_METER_DISPLAY := 26389, NEXT_SCHDL_MAINTENANCE := 2, MAINTENANCE_ALARM := 1);
   _35_JUMP_LEG_RUNNING : BOOL := 1;
   _35AUTO : ALIAS FOR B9[35].4;
   _35HAND : ALIAS FOR B9[35].3;
   _35M : ALIAS FOR O25[10].13;
   _35MB : ALIAS FOR B9[35].2;
   _35STB : ALIAS FOR B9[35].0;
   _35STPB : ALIAS FOR B9[35].1;
   _35Y : ALIAS FOR I25[2].13;
   _36_FREQ_IN : ALIAS FOR N7[1];
   _36_FREQ_OU : ALIAS FOR N7[3];
   _36_SET_SPD : ALIAS FOR N7[2];
   _36_TANK_41_AUGER_HM : HOUR_METER := (HR_METER_DISPLAY := 2995, MAINTENANCE_ALARM := 1);
   _36_VFD_TO : ALIAS FOR N180[0];
   _36M : ALIAS FOR O25[8].0;
   _36MAI : ALIAS FOR O25[25].0;
   _36RAUTO : ALIAS FOR B9[36].4;
   _36RHAND : ALIAS FOR B9[36].3;
   _36RMB : ALIAS FOR B9[36].2;
   _36RSTB : ALIAS FOR B9[36].0;
   _36RSTPB : ALIAS FOR B9[36].1;
   _36RY : ALIAS FOR I25[16].0;
   _36Y : ALIAS FOR I25[0].0;
   _3_LOWER_TANK_CONVAYOR_24TO26_HM : HOUR_METER := (HR_METER_DISPLAY := 1012, NEXT_SCHDL_MAINTENANCE := 2, MAINTENANCE_ALARM := 1);
   _3_LOWER_TANK_CONVAYOR_24TO26_RUNNING : BOOL;
   _3_LS_TO_5 : ALIAS FOR I25[4].8;
   _3_LS_TO_6 : ALIAS FOR I25[4].9;
   _3_TO_BC5_S : ALIAS FOR O25[11].12;
   _3_TO_BC6_S : ALIAS FOR O25[11].13;
   _3AUTO : ALIAS FOR B9[3].4;
   _3HAND : ALIAS FOR B9[3].3;
   _3M : ALIAS FOR O25[10].0;
   _3MB : ALIAS FOR B9[3].2;
   _3STB : ALIAS FOR B9[3].0;
   _3STPB : ALIAS FOR B9[3].1;
   _3Y : ALIAS FOR I25[2].0;
   _41_GATE_PO : ALIAS FOR I18[0];
   _41_GATE_PO1 : ALIAS FOR N14[41];
   _42_GATE_PO : ALIAS FOR I18[1];
   _42_GATE_PO1 : ALIAS FOR N14[42];
   _42_LOWER_SCREENINGS_DRAG_HM : HOUR_METER := (MOTOR_RUNNING_INPUT_1 := 1, HR_METER_DISPLAY := 27637, MAINTENANCE_ALARM := 1);
   _42AUTO : ALIAS FOR B9[42].4;
   _42HAND : ALIAS FOR B9[42].3;
   _42M : ALIAS FOR O25[11].1;
   _42MB : ALIAS FOR B9[42].2;
   _42STB : ALIAS FOR B9[42].0;
   _42STPB : ALIAS FOR B9[42].1;
   _42Y : ALIAS FOR I25[3].1;
   _43_ACC_WEI : ALIAS FOR C5[1].ACC;
   _43_BINDICA : ALIAS FOR B9[43].5;
   _43_RESET_C : ALIAS FOR B9[43].6;
   _43_SCREEN : ALIAS FOR C5[1];
   _43_SCREENI : ALIAS FOR I7.14;
   _43_SCREENINGS_LEG_HM : HOUR_METER := (MOTOR_RUNNING_INPUT_1 := 1, HR_METER_DISPLAY := 27656, NEXT_SCHDL_MAINTENANCE := 2, MAINTENANCE_ALARM := 1);
   _43_SCREENINGS_LEG_RUNNING : BOOL := 1;
   _43_WEIGHT : ALIAS FOR N7[0];
   _43AUTO : ALIAS FOR B9[43].4;
   _43HAND : ALIAS FOR B9[43].3;
   _43M : ALIAS FOR O25[10].14;